
screen "4. VFD 10 - 13" 1280x800, template "Main_Template"
   on GenerateScreen: SetTag("animation_page", 4)
   Bar "Bar_1" at 206,213 size 88x440; MinimumValue 0; MaximumValue 50
      ProcessValue <- "speedActual_address_10"
   Button "Button_7" at 35,514 size 150x62; TextOff '+'
      on Press: function_b14e0dd5("increaseSpeed_address_10", 0)
      Appearance <- "statusIncrease_address_10"
   Button "Button_8" at 35,591 size 150x62; TextOff '-'
      on Press: function_b14e0dd5("decreaseSpeed_address_10", 0)
      Appearance <- "statusDecrease_address_10"
   TextField "Text field_20" at 35,428 size 150x62; Text 'Hz'
   IOField "I/O field_1" at 37,430 size 98x57; FormatPattern 99.99
      ProcessValue <- "speedActual_address_10"
   TextField "Text field_14" at 28,133 size 207x62; Text 'Gauge Roll 3rd Set'
   TextField "Text field_26" at 35,228 size 150x62; Text 'Hz'
   TextField "Text field_32" at 35,328 size 150x62; Text 'Hz'
   IOField "I/O field_2" at 39,231 size 98x57; FormatPattern 99.99
      ProcessValue <- "speedReff_singleSync_address_10"
   TextField "Text field_1" at 35,400 size 115x27; Text 'Actual Speed'
   TextField "Text field_2" at 35,302 size 144x27; Text 'Reff Speed Sync'
   TextField "Text field_3" at 35,200 size 155x27; Text 'Reff Speed Single'
   TextField "Text field_4" at 36,661 size 149x45; Text 'VFD 10'
      Appearance <- "Running_Motor Addres_10"
   Bar "Bar_2" at 518,213 size 88x440; MinimumValue 0; MaximumValue 50
      ProcessValue <- "speedActual_address_11"
   Button "Button_2" at 347,514 size 150x62; TextOff '+'
      on Press: function_b14e0dd5("increaseSpeed_address_11", 0)
      Appearance <- "statusIncrease_address_11"
   Button "Button_3" at 347,591 size 150x62; TextOff '-'
      on Press: function_b14e0dd5("decreaseSpeed_address_11", 0)
      Appearance <- "statusDecrease_address_11"
   TextField "Text field_5" at 347,428 size 150x62; Text 'Hz'
   IOField "I/O field_3" at 349,430 size 98x57; FormatPattern 99.99
      ProcessValue <- "speedActual_address_11"
   TextField "Text field_6" at 340,133 size 207x62; Text 'Conveyor of Gauge Roll 3rd Set'
   TextField "Text field_7" at 347,228 size 150x62; Text 'Hz'
   TextField "Text field_8" at 347,328 size 150x62; Text 'Hz'
   IOField "I/O field_4" at 351,231 size 98x57; FormatPattern 99.99
      ProcessValue <- "speedReff_singleSync_address_11"
   TextField "Text field_9" at 347,400 size 115x27; Text 'Actual Speed'
   TextField "Text field_10" at 347,302 size 144x27; Text 'Reff Speed Sync'
   TextField "Text field_11" at 347,200 size 155x27; Text 'Reff Speed Single'
   TextField "Text field_12" at 348,661 size 149x45; Text 'VFD 11'
      Appearance <- "Running_Motor Addres_11"
   Bar "Bar_3" at 830,213 size 88x440; MinimumValue 0; MaximumValue 50
      ProcessValue <- "speedActual_address_12"
   Button "Button_4" at 659,514 size 150x62; TextOff '+'
      on Press: function_b14e0dd5("increaseSpeed_address_12", 0)
      Appearance <- "statusIncrease_address_12"
   Button "Button_5" at 659,591 size 150x62; TextOff '-'
      on Press: function_b14e0dd5("decreaseSpeed_address_12", 0)
      Appearance <- "statusDecrease_address_12"
   TextField "Text field_13" at 659,428 size 150x62; Text 'Hz'
   IOField "I/O field_5" at 661,430 size 98x57; FormatPattern 99.99
      ProcessValue <- "speedActual_address_12"
   TextField "Text field_15" at 652,133 size 207x62; Text 'Passing Conveyor of Rotary Mould'
   TextField "Text field_16" at 659,228 size 150x62; Text 'Hz'
   TextField "Text field_17" at 659,328 size 150x62; Text 'Hz'
   IOField "I/O field_6" at 663,231 size 98x57; FormatPattern 99.99
      ProcessValue <- "speedReff_singleSync_address_12"
   TextField "Text field_18" at 659,400 size 115x27; Text 'Actual Speed'
   TextField "Text field_19" at 659,302 size 144x27; Text 'Reff Speed Sync'
   TextField "Text field_21" at 659,200 size 155x27; Text 'Reff Speed Single'
   TextField "Text field_22" at 660,661 size 149x45; Text 'VFD 12'
      Appearance <- "Running_Motor Addres_12"
   Bar "Bar_4" at 1142,213 size 88x440; MinimumValue 0; MaximumValue 50
      ProcessValue <- "speedActual_address_13"
   Button "Button_6" at 971,514 size 150x62; TextOff '+'
      on Press: function_b14e0dd5("increaseSpeed_address_13", 0)
      Appearance <- "statusIncrease_address_13"
   Button "Button_9" at 971,591 size 150x62; TextOff '-'
      on Press: function_b14e0dd5("decreaseSpeed_address_13", 0)
      Appearance <- "statusDecrease_address_13"
   TextField "Text field_23" at 971,428 size 150x62; Text 'Hz'
   IOField "I/O field_7" at 973,430 size 98x57; FormatPattern 99.99
      ProcessValue <- "speedActual_address_13"
   TextField "Text field_24" at 964,133 size 207x62; Text 'Conveyor of Rotary Moulder'
   TextField "Text field_25" at 971,228 size 150x62; Text 'Hz'
   TextField "Text field_27" at 971,328 size 150x62; Text 'Hz'
   IOField "I/O field_8" at 975,231 size 98x57; FormatPattern 99.99
      ProcessValue <- "speedReff_singleSync_address_13"
   TextField "Text field_28" at 971,400 size 115x27; Text 'Actual Speed'
   TextField "Text field_29" at 971,302 size 144x27; Text 'Reff Speed Sync'
   TextField "Text field_30" at 971,200 size 155x27; Text 'Reff Speed Single'
   TextField "Text field_31" at 972,661 size 149x45; Text 'VFD 13'
      Appearance <- "Running_Motor Addres_13"
   IOField "I/O field_14" at 349,330 size 98x57; FormatPattern 99.99
      ProcessValue <- "speedReff_NOT_singleSync_address_11"
   IOField "I/O field_9" at 661,330 size 98x57; FormatPattern 99.99
      ProcessValue <- "speedReff_NOT_singleSync_address_12"
   IOField "I/O field_10" at 973,330 size 98x57; FormatPattern 99.99
      ProcessValue <- "speedReff_NOT_singleSync_address_13"
   SymbolicIOField "Symbolic I/O field_2" at 550,133 size 77x62; TextOn '1'; TextOff '0'; TextList "Mode_Syncron"
      Appearance <- "Syncron_2"
      ProcessValue <- "Syncron_2"
   SymbolicIOField "Symbolic I/O field_3" at 862,133 size 77x62; TextOn '1'; TextOff '0'; TextList "Mode_Syncron"
      Appearance <- "Syncron_2"
      ProcessValue <- "Syncron_2"
   SymbolicIOField "Symbolic I/O field_4" at 1174,133 size 77x62; TextOn '1'; TextOff '0'; TextList "Mode_Syncron"
      Appearance <- "Syncron_1"
      ProcessValue <- "Syncron_1"
   IOField "I/O field_11" at 37,330 size 98x57; FormatPattern 99.99
      ProcessValue <- "speedReff_NOT_singleSync_address_10"
   SymbolicIOField "Symbolic I/O field_1" at 238,133 size 77x62; TextOn '1'; TextOff '0'; TextList "Mode_Syncron"
      Appearance <- "Syncron_2"
      ProcessValue <- "Syncron_2"
   Button "Button_1" at 0,721 size 160x79; TextOff 'MAIN'
      on Click: ActivateScreen("1. MAIN", 0)
      Appearance <- "animation_page"
   Button "Button_10" at 160,721 size 160x79; TextOff 'VFD 2 - 5'
      on Click: ActivateScreen("2. VFD 2 - 5", 0)
      Appearance <- "animation_page"
   Button "Button_11" at 320,721 size 160x79; TextOff 'VFD 6 - 9'
      on Click: ActivateScreen("3. VFD 6 - 9", 0)
      Appearance <- "animation_page"
   Button "Button_12" at 480,721 size 160x79; TextOff 'VFD 10 - 13'
      on Click: ActivateScreen("4. VFD 10 - 13", 0)
      Appearance <- "animation_page"
   Button "Button_13" at 640,721 size 160x79; TextOff 'VFD 14 - 17'
      on Click: ActivateScreen("5. VFD 14 - 17", 0)
      Appearance <- "animation_page"
   Button "Button_14" at 800,721 size 160x79; TextOff 'VFD 18 - 21'
      on Click: ActivateScreen("6. VFD 18 - 21", 0)
      Appearance <- "animation_page"
   Button "Button_15" at 960,721 size 160x79; TextOff 'VFD 22 - 23'
      on Click: ActivateScreen("7. VFD 22 - 23", 0)
      Appearance <- "animation_page"
   Button "Button_16" at 1120,721 size 160x79; TextOff 'Alarm'
      on Click: ActivateScreen("8. ALARM", 0)
      Appearance <- "animation_page"
   TextField "Text field_34" at 0,64 size 331x50; Text 'MOTOR CONTROL SPEED'
   Softkey "Softkey_F1" at 0,0 size 0x0
      on KeyDown: ActivateScreen("1. MAIN", 0)
   Softkey "Softkey_F2" at 0,0 size 0x0
      on KeyDown: ActivateScreen("2. VFD 2 - 5", 0)
   Softkey "Softkey_F3" at 0,0 size 0x0
      on KeyDown: ActivateScreen("3. VFD 6 - 9", 0)
   Softkey "Softkey_F4" at 0,0 size 0x0
      on KeyDown: ActivateScreen("4. VFD 10 - 13", 0)
   Softkey "Softkey_F5" at 0,0 size 0x0
      on KeyDown: ActivateScreen("5. VFD 14 - 17", 0)
   Softkey "Softkey_F6" at 0,0 size 0x0
      on KeyDown: ActivateScreen("6. VFD 18 - 21", 0)
   Softkey "Softkey_F7" at 0,0 size 0x0
      on KeyDown: ActivateScreen("7. VFD 22 - 23", 0)
   Softkey "Softkey_F8" at 0,0 size 0x0
      on KeyDown: ActivateScreen("8. ALARM", 0)
   Softkey "Softkey_F9" at 0,0 size 0x0
      on KeyDown: ActivateScreen("9. VFD PROFIBUS", 0)
   Softkey "Softkey_F10" at 0,0 size 0x0
      on KeyDown: ActivateScreen("10. SETTINGS", 0)

screen "5. VFD 14 - 17" 1280x800, template "Main_Template"
   on GenerateScreen: SetTag("animation_page", 5)
   Bar "Bar_1" at 206,213 size 88x440; MinimumValue 0; MaximumValue 50
      ProcessValue <- "speedActual_address_14"
   Button "Button_7" at 35,514 size 150x62; TextOff '+'
      on Press: function_b14e0dd5("increaseSpeed_address_14", 0)
      Appearance <- "statusIncrease_address_14"
   Button "Button_8" at 35,591 size 150x62; TextOff '-'
      on Press: function_b14e0dd5("decreaseSpeed_address_14", 0)
      Appearance <- "statusDecrease_address_14"
   TextField "Text field_20" at 35,428 size 150x62; Text 'Hz'
   IOField "I/O field_1" at 37,430 size 98x57; FormatPattern 99.99
      ProcessValue <- "speedActual_address_14"
   TextField "Text field_14" at 28,133 size 207x62; Text 'Drive of Mould'
   TextField "Text field_26" at 35,228 size 150x62; Text 'Hz'
   TextField "Text field_32" at 35,328 size 150x62; Text 'Hz'
   IOField "I/O field_2" at 39,231 size 98x57; FormatPattern 99.99
      ProcessValue <- "speedReff_singleSync_address_14"
   TextField "Text field_1" at 35,400 size 115x27; Text 'Actual Speed'
   TextField "Text field_2" at 35,302 size 144x27; Text 'Reff Speed Sync'
   TextField "Text field_3" at 35,200 size 155x27; Text 'Reff Speed Single'
   TextField "Text field_4" at 36,661 size 149x45; Text 'VFD 14'
      Appearance <- "Running_Motor Addres_14"
   Bar "Bar_2" at 518,213 size 88x440; MinimumValue 0; MaximumValue 50
      ProcessValue <- "speedActual_address_15"
   Button "Button_2" at 347,514 size 150x62; TextOff '+'
      on Press: function_b14e0dd5("increaseSpeed_address_15", 0)
      Appearance <- "statusIncrease_address_15"
   Button "Button_3" at 347,591 size 150x62; TextOff '-'
      on Press: function_b14e0dd5("decreaseSpeed_address_15", 0)
      Appearance <- "statusDecrease_address_15"
   TextField "Text field_5" at 347,428 size 150x62; Text 'Hz'
   IOField "I/O field_3" at 349,430 size 98x57; FormatPattern 99.99
      ProcessValue <- "speedActual_address_15"
   TextField "Text field_6" at 340,133 size 207x62; Text 'Forcing Roll'
   TextField "Text field_7" at 347,228 size 150x62; Text 'Hz'
   TextField "Text field_8" at 347,328 size 150x62; Text 'Hz'
   IOField "I/O field_4" at 351,231 size 98x57; FormatPattern 99.99
      ProcessValue <- "speedReff_singleSync_address_15"
   TextField "Text field_9" at 347,400 size 115x27; Text 'Actual Speed'
   TextField "Text field_10" at 347,302 size 144x27; Text 'Reff Speed Sync'
   TextField "Text field_11" at 347,200 size 155x27; Text 'Reff Speed Single'
   TextField "Text field_12" at 348,661 size 149x45; Text 'VFD 15'
      Appearance <- "Running_Motor Addres_15"
   Bar "Bar_3" at 830,213 size 88x440; MinimumValue 0; MaximumValue 50
      ProcessValue <- "speedActual_address_16"
   Button "Button_4" at 659,514 size 150x62; TextOff '+'
      on Press: function_b14e0dd5("increaseSpeed_address_16", 0)
      Appearance <- "statusIncrease_address_16"
   Button "Button_5" at 659,591 size 150x62; TextOff '-'
      on Press: function_b14e0dd5("decreaseSpeed_address_16", 0)
      Appearance <- "statusDecrease_address_16"
   TextField "Text field_13" at 659,428 size 150x62; Text 'Hz'
   IOField "I/O field_5" at 661,430 size 98x57; FormatPattern 99.99
      ProcessValue <- "speedActual_address_16"
   TextField "Text field_15" at 652,133 size 207x62; Text 'Mould of Rotary Cutter'
   TextField "Text field_16" at 659,228 size 150x62; Text 'Hz'
   TextField "Text field_17" at 659,328 size 150x62; Text 'Hz'
   IOField "I/O field_6" at 663,231 size 98x57; FormatPattern 99.99
      ProcessValue <- "speedReff_singleSync_address_16"
   TextField "Text field_18" at 659,400 size 115x27; Text 'Actual Speed'
   TextField "Text field_19" at 659,302 size 144x27; Text 'Reff Speed Sync'
   TextField "Text field_21" at 659,200 size 155x27; Text 'Reff Speed Single'
   TextField "Text field_22" at 660,661 size 149x45; Text 'VFD 16'
      Appearance <- "Running_Motor Addres_16"
   Bar "Bar_4" at 1142,213 size 88x440; MinimumValue 0; MaximumValue 50
      ProcessValue <- "speedActual_address_17"
   Button "Button_6" at 971,514 size 150x62; TextOff '+'
      on Press: function_b14e0dd5("increaseSpeed_address_17", 0)
      Appearance <- "statusIncrease_address_17"
   Button "Button_9" at 971,591 size 150x62; TextOff '-'
      on Press: function_b14e0dd5("decreaseSpeed_address_17", 0)
      Appearance <- "statusDecrease_address_17"
   TextField "Text field_23" at 971,428 size 150x62; Text 'Hz'
   IOField "I/O field_7" at 973,430 size 98x57; FormatPattern 99.99
      ProcessValue <- "speedActual_address_17"
   TextField "Text field_24" at 964,133 size 207x62; Text 'Conveyor for Rotary Cutter'
   TextField "Text field_25" at 971,228 size 150x62; Text 'Hz'
   TextField "Text field_27" at 971,328 size 150x62; Text 'Hz'
   IOField "I/O field_8" at 975,231 size 98x57; FormatPattern 99.99
      ProcessValue <- "speedReff_singleSync_address_17"
   TextField "Text field_28" at 971,400 size 115x27; Text 'Actual Speed'
   TextField "Text field_29" at 971,302 size 144x27; Text 'Reff Speed Sync'
   TextField "Text field_30" at 971,200 size 155x27; Text 'Reff Speed Single'
   TextField "Text field_31" at 972,661 size 149x45; Text 'VFD 17'
      Appearance <- "Running_Motor Addres_17"
   IOField "I/O field_14" at 349,330 size 98x57; FormatPattern 99.99
      ProcessValue <- "speedReff_NOT_singleSync_address_15"
   IOField "I/O field_9" at 661,330 size 98x57; FormatPattern 99.99
      ProcessValue <- "speedReff_NOT_singleSync_address_16"
   IOField "I/O field_10" at 973,330 size 98x57; FormatPattern 99.99
      ProcessValue <- "speedReff_NOT_singleSync_address_17"
   SymbolicIOField "Symbolic I/O field_2" at 550,133 size 77x62; TextOn '1'; TextOff '0'; TextList "Mode_Syncron"
      Appearance <- "Syncron_1"
      ProcessValue <- "Syncron_1"
   SymbolicIOField "Symbolic I/O field_3" at 862,133 size 77x62; TextOn '1'; TextOff '0'; TextList "Mode_Syncron"
      Appearance <- "Syncron_2"
      ProcessValue <- "Syncron_2"
   SymbolicIOField "Symbolic I/O field_4" at 1174,133 size 77x62; TextOn '1'; TextOff '0'; TextList "Mode_Syncron"
      Appearance <- "Syncron_3"
      ProcessValue <- "Syncron_3"
   IOField "I/O field_11" at 37,330 size 98x57; FormatPattern 99.99
      ProcessValue <- "speedReff_NOT_singleSync_address_14"
   SymbolicIOField "Symbolic I/O field_1" at 238,133 size 77x62; TextOn '1'; TextOff '0'; TextList "Mode_Syncron"
      Appearance <- "Syncron_1"
      ProcessValue <- "Syncron_1"
   Button "Button_1" at 0,721 size 160x79; TextOff 'MAIN'
      on Click: ActivateScreen("1. MAIN", 0)
      Appearance <- "animation_page"
   Button "Button_10" at 160,721 size 160x79; TextOff 'VFD 2 - 5'
      on Click: ActivateScreen("2. VFD 2 - 5", 0)
      Appearance <- "animation_page"
   Button "Button_11" at 320,721 size 160x79; TextOff 'VFD 6 - 9'
      on Click: ActivateScreen("3. VFD 6 - 9", 0)
      Appearance <- "animation_page"
   Button "Button_12" at 480,721 size 160x79; TextOff 'VFD 10 - 13'
      on Click: ActivateScreen("4. VFD 10 - 13", 0)
      Appearance <- "animation_page"
   Button "Button_13" at 640,721 size 160x79; TextOff 'VFD 14 - 17'
      on Click: ActivateScreen("5. VFD 14 - 17", 0)
      Appearance <- "animation_page"
   Button "Button_14" at 800,721 size 160x79; TextOff 'VFD 18 - 21'
      on Click: ActivateScreen("6. VFD 18 - 21", 0)
      Appearance <- "animation_page"
   Button "Button_15" at 960,721 size 160x79; TextOff 'VFD 22 - 23'
      on Click: ActivateScreen("7. VFD 22 - 23", 0)
      Appearance <- "animation_page"
   Button "Button_16" at 1120,721 size 160x79; TextOff 'Alarm'
      on Click: ActivateScreen("8. ALARM", 0)
      Appearance <- "animation_page"
   TextField "Text field_34" at 0,64 size 331x50; Text 'MOTOR CONTROL SPEED'
   Softkey "Softkey_F5" at 0,0 size 0x0
      on KeyDown: ActivateScreen("5. VFD 14 - 17", 0)
   Softkey "Softkey_F1" at 0,0 size 0x0
      on KeyDown: ActivateScreen("1. MAIN", 0)
   Softkey "Softkey_F2" at 0,0 size 0x0
      on KeyDown: ActivateScreen("2. VFD 2 - 5", 0)
   Softkey "Softkey_F3" at 0,0 size 0x0
      on KeyDown: ActivateScreen("3. VFD 6 - 9", 0)
   Softkey "Softkey_F4" at 0,0 size 0x0
      on KeyDown: ActivateScreen("4. VFD 10 - 13", 0)
   Softkey "Softkey_F6" at 0,0 size 0x0
      on KeyDown: ActivateScreen("6. VFD 18 - 21", 0)
   Softkey "Softkey_F7" at 0,0 size 0x0
      on KeyDown: ActivateScreen("7. VFD 22 - 23", 0)
   Softkey "Softkey_F8" at 0,0 size 0x0
      on KeyDown: ActivateScreen("8. ALARM", 0)
   Softkey "Softkey_F9" at 0,0 size 0x0
      on KeyDown: ActivateScreen("9. VFD PROFIBUS", 0)
   Softkey "Softkey_F10" at 0,0 size 0x0
      on KeyDown: ActivateScreen("10. SETTINGS", 0)

screen "6. VFD 18 - 21" 1280x800, template "Main_Template"
   on GenerateScreen: SetTag("animation_page", 6)
   Bar "Bar_1" at 206,213 size 88x440; MinimumValue 0; MaximumValue 50
      ProcessValue <- "speedActual_address_18"
   Button "Button_7" at 35,514 size 150x62; TextOff '+'
      on Press: function_b14e0dd5("increaseSpeed_address_18", 0)
      Appearance <- "statusIncrease_address_18"
   Button "Button_8" at 35,591 size 150x62; TextOff '-'
      on Press: function_b14e0dd5("decreaseSpeed_address_18", 0)
      Appearance <- "statusDecrease_address_18"
   TextField "Text field_20" at 35,428 size 150x62; Text 'Hz'
   IOField "I/O field_1" at 37,430 size 98x57; FormatPattern 99.99
      ProcessValue <- "speedActual_address_18"
   TextField "Text field_14" at 28,133 size 207x62; Text 'Dough Feed for Rotary Moulder'
   TextField "Text field_26" at 35,228 size 150x62; Text 'Hz'
   TextField "Text field_32" at 35,328 size 150x62; Text 'Hz'
   IOField "I/O field_2" at 39,231 size 98x57; FormatPattern 99.99
      ProcessValue <- "speedReff_singleSync_address_18"
   TextField "Text field_1" at 35,400 size 115x27; Text 'Actual Speed'
   TextField "Text field_2" at 35,302 size 144x27; Text 'Reff Speed Sync'
   TextField "Text field_3" at 35,200 size 155x27; Text 'Reff Speed Single'
   TextField "Text field_4" at 36,661 size 149x45; Text 'VFD 18'
      Appearance <- "Running_Motor Addres_18"
   Bar "Bar_2" at 518,213 size 88x440; MinimumValue 0; MaximumValue 50
      ProcessValue <- "speedActual_address_19"
   Button "Button_2" at 347,514 size 150x62; TextOff '+'
      on Press: function_b14e0dd5("increaseSpeed_address_19", 0)
      Appearance <- "statusIncrease_address_19"
   Button "Button_3" at 347,591 size 150x62; TextOff '-'
      on Press: function_b14e0dd5("decreaseSpeed_address_19", 0)
      Appearance <- "statusDecrease_address_19"
   TextField "Text field_5" at 347,428 size 150x62; Text 'Hz'
   IOField "I/O field_3" at 349,430 size 98x57; FormatPattern 99.99
      ProcessValue <- "speedActual_address_19"
   TextField "Text field_6" at 340,133 size 207x62; Text 'Conveyor of Scrapt Lift Passing'
   TextField "Text field_7" at 347,228 size 150x62; Text 'Hz'
   TextField "Text field_8" at 347,328 size 150x62; Text 'Hz'
   IOField "I/O field_4" at 351,231 size 98x57; FormatPattern 99.99
      ProcessValue <- "speedReff_singleSync_address_19"
   TextField "Text field_9" at 347,400 size 115x27; Text 'Actual Speed'
   TextField "Text field_10" at 347,302 size 144x27; Text 'Reff Speed Sync'
   TextField "Text field_11" at 347,200 size 155x27; Text 'Reff Speed Single'
   TextField "Text field_12" at 348,661 size 149x45; Text 'VFD 19'
      Appearance <- "Running_Motor Addres_19"
   Bar "Bar_3" at 830,213 size 88x440; MinimumValue 0; MaximumValue 50
      ProcessValue <- "speedActual_address_20"
   Button "Button_4" at 659,514 size 150x62; TextOff '+'
      on Press: function_b14e0dd5("increaseSpeed_address_20", 0)
      Appearance <- "statusIncrease_address_20"
   Button "Button_5" at 659,591 size 150x62; TextOff '-'
      on Press: function_b14e0dd5("decreaseSpeed_address_20", 0)
      Appearance <- "statusDecrease_address_20"
   TextField "Text field_13" at 659,428 size 150x62; Text 'Hz'
   IOField "I/O field_5" at 661,430 size 98x57; FormatPattern 99.99
      ProcessValue <- "speedActual_address_20"
   TextField "Text field_15" at 652,133 size 207x62; Text 'Conveyor of Salt Sprinkler'
   TextField "Text field_16" at 659,228 size 150x62; Text 'Hz'
   TextField "Text field_17" at 659,328 size 150x62; Text 'Hz'
   IOField "I/O field_6" at 663,231 size 98x57; FormatPattern 99.99
      ProcessValue <- "speedReff_singleSync_address_20"
   TextField "Text field_18" at 659,400 size 115x27; Text 'Actual Speed'
   TextField "Text field_19" at 659,302 size 144x27; Text 'Reff Speed Sync'
   TextField "Text field_21" at 659,200 size 155x27; Text 'Reff Speed Single'
   TextField "Text field_22" at 660,661 size 149x45; Text 'VFD 20'
      Appearance <- "Running_Motor Addres_20"
   Bar "Bar_4" at 1142,213 size 88x440; MinimumValue 0; MaximumValue 50
      ProcessValue <- "speedActual_address_21"
   Button "Button_6" at 971,514 size 150x62; TextOff '+'
      on Press: function_b14e0dd5("increaseSpeed_address_21", 0)
      Appearance <- "statusIncrease_address_21"
   Button "Button_9" at 971,591 size 150x62; TextOff '-'
      on Press: function_b14e0dd5("decreaseSpeed_address_21", 0)
      Appearance <- "statusDecrease_address_21"
   TextField "Text field_23" at 971,428 size 150x62; Text 'Hz'
   IOField "I/O field_7" at 973,430 size 98x57; FormatPattern 99.99
      ProcessValue <- "speedActual_address_21"
   TextField "Text field_24" at 964,133 size 207x62; Text 'Recovery Conveyor of Salt Sprinkler'
   TextField "Text field_25" at 971,228 size 150x62; Text 'Hz'
   TextField "Text field_27" at 971,328 size 150x62; Text 'Hz'
   IOField "I/O field_8" at 975,231 size 98x57; FormatPattern 99.99
      ProcessValue <- "speedReff_singleSync_address_21"
   TextField "Text field_28" at 971,400 size 115x27; Text 'Actual Speed'
   TextField "Text field_29" at 971,302 size 144x27; Text 'Reff Speed Sync'
   TextField "Text field_30" at 971,200 size 155x27; Text 'Reff Speed Single'
   TextField "Text field_31" at 972,661 size 149x45; Text 'VFD 21'
      Appearance <- "Running_Motor Addres_21"
   IOField "I/O field_14" at 349,330 size 98x57; FormatPattern 99.99
      ProcessValue <- "speedReff_NOT_singleSync_address_19"
   IOField "I/O field_9" at 661,330 size 98x57; FormatPattern 99.99
      ProcessValue <- "speedReff_NOT_singleSync_address_20"
   IOField "I/O field_10" at 973,330 size 98x57; FormatPattern 99.99
      ProcessValue <- "speedReff_NOT_singleSync_address_21"
   SymbolicIOField "Symbolic I/O field_2" at 550,133 size 77x62; TextOn '1'; TextOff '0'; TextList "Mode_Syncron"
      Appearance <- "Syncron_3"
      ProcessValue <- "Syncron_3"
   SymbolicIOField "Symbolic I/O field_4" at 1174,133 size 77x62; TextOn '1'; TextOff '0'; TextList "Mode_Syncron"
      Appearance <- "Syncron_3"
      ProcessValue <- "Syncron_3"
   IOField "I/O field_11" at 37,330 size 98x57; FormatPattern 99.99
      ProcessValue <- "speedReff_NOT_singleSync_address_18"
   TextField "Text field_33" at 238,133 size 76x62; Text 'Single'
   TextField "Text field_35" at 863,133 size 76x62; Text 'Single'
   Button "Button_1" at 0,721 size 160x79; TextOff 'MAIN'
      on Click: ActivateScreen("1. MAIN", 0)
      Appearance <- "animation_page"
   Button "Button_10" at 160,721 size 160x79; TextOff 'VFD 2 - 5'
      on Click: ActivateScreen("2. VFD 2 - 5", 0)
      Appearance <- "animation_page"
   Button "Button_11" at 320,721 size 160x79; TextOff 'VFD 6 - 9'
      on Click: ActivateScreen("3. VFD 6 - 9", 0)
      Appearance <- "animation_page"
   Button "Button_12" at 480,721 size 160x79; TextOff 'VFD 10 - 13'
      on Click: ActivateScreen("4. VFD 10 - 13", 0)
      Appearance <- "animation_page"
   Button "Button_13" at 640,721 size 160x79; TextOff 'VFD 14 - 17'
      on Click: ActivateScreen("5. VFD 14 - 17", 0)
      Appearance <- "animation_page"
   Button "Button_14" at 800,721 size 160x79; TextOff 'VFD 18 - 21'
      on Click: ActivateScreen("6. VFD 18 - 21", 0)
      Appearance <- "animation_page"
   Button "Button_15" at 960,721 size 160x79; TextOff 'VFD 22 - 23'
      on Click: ActivateScreen("7. VFD 22 - 23", 0)
      Appearance <- "animation_page"
   Button "Button_16" at 1120,721 size 160x79; TextOff 'Alarm'
      on Click: ActivateScreen("8. ALARM", 0)
      Appearance <- "animation_page"
   TextField "Text field_34" at 0,64 size 331x50; Text 'MOTOR CONTROL SPEED'
   Softkey "Softkey_F5" at 0,0 size 0x0
      on KeyDown: ActivateScreen("5. VFD 14 - 17", 0)
   Softkey "Softkey_F1" at 0,0 size 0x0
      on KeyDown: ActivateScreen("1. MAIN", 0)
   Softkey "Softkey_F2" at 0,0 size 0x0
      on KeyDown: ActivateScreen("2. VFD 2 - 5", 0)
   Softkey "Softkey_F3" at 0,0 size 0x0
      on KeyDown: ActivateScreen("3. VFD 6 - 9", 0)
   Softkey "Softkey_F4" at 0,0 size 0x0
      on KeyDown: ActivateScreen("4. VFD 10 - 13", 0)
   Softkey "Softkey_F6" at 0,0 size 0x0
      on KeyDown: ActivateScreen("6. VFD 18 - 21", 0)
   Softkey "Softkey_F7" at 0,0 size 0x0
      on KeyDown: ActivateScreen("7. VFD 22 - 23", 0)
   Softkey "Softkey_F8" at 0,0 size 0x0
      on KeyDown: ActivateScreen("8. ALARM", 0)
   Softkey "Softkey_F9" at 0,0 size 0x0
      on KeyDown: ActivateScreen("9. VFD PROFIBUS", 0)
   Softkey "Softkey_F10" at 0,0 size 0x0
      on KeyDown: ActivateScreen("10. SETTINGS", 0)

screen "7. VFD 22 - 23" 1280x800, template "Main_Template"
   on GenerateScreen: SetTag("animation_page", 7)
   Bar "Bar_1" at 206,213 size 88x440; MinimumValue 0; MaximumValue 50
      ProcessValue <- "speedActual_address_22"
   Button "Button_7" at 35,514 size 150x62; TextOff '+'
      on Press: function_b14e0dd5("increaseSpeed_address_22", 0)
      Appearance <- "statusIncrease_address_22"
   Button "Button_8" at 35,591 size 150x62; TextOff '-'
      on Press: function_b14e0dd5("decreaseSpeed_address_22", 0)
      Appearance <- "statusDecrease_address_22"
   TextField "Text field_20" at 35,428 size 150x62; Text 'Hz'
   IOField "I/O field_1" at 37,430 size 98x57; FormatPattern 99.99
      ProcessValue <- "speedActual_address_22"
   TextField "Text field_14" at 28,133 size 207x62; Text 'Conveyor Swivel Panner'
   TextField "Text field_26" at 35,228 size 150x62; Text 'Hz'
   TextField "Text field_32" at 35,328 size 150x62; Text 'Hz'
   IOField "I/O field_2" at 39,231 size 98x57; FormatPattern 99.99
      ProcessValue <- "speedReff_singleSync_address_22"
   TextField "Text field_1" at 35,400 size 115x27; Text 'Actual Speed'
   TextField "Text field_2" at 35,302 size 144x27; Text 'Reff Speed Sync'
   TextField "Text field_3" at 35,200 size 155x27; Text 'Reff Speed Single'
   TextField "Text field_4" at 36,661 size 149x45; Text 'VFD 22'
      Appearance <- "Running_Motor Addres_22"
   Bar "Bar_2" at 518,213 size 88x440; MinimumValue 0; MaximumValue 50
      ProcessValue <- "speedActual_address_23"
   Button "Button_2" at 347,514 size 150x62; TextOff '+'
      on Press: function_b14e0dd5("increaseSpeed_address_23", 0)
      Appearance <- "statusIncrease_address_23"
   Button "Button_3" at 347,591 size 150x62; TextOff '-'
      on Press: function_b14e0dd5("decreaseSpeed_address_23", 0)
      Appearance <- "statusDecrease_address_23"
   TextField "Text field_5" at 347,428 size 150x62; Text 'Hz'
   IOField "I/O field_3" at 349,430 size 98x57; FormatPattern 99.99
      ProcessValue <- "speedActual_address_23"
   TextField "Text field_6" at 340,133 size 207x62; Text 'Side Return VFD 23 for 4 Motor'
   TextField "Text field_7" at 347,228 size 150x62; Text 'Hz'
   TextField "Text field_8" at 347,328 size 150x62; Text 'Hz'
   IOField "I/O field_4" at 351,231 size 98x57; FormatPattern 99.99
      ProcessValue <- "speedReff_singleSync_address_23"
   TextField "Text field_9" at 347,400 size 115x27; Text 'Actual Speed'
   TextField "Text field_10" at 347,302 size 144x27; Text 'Reff Speed Sync'
   TextField "Text field_11" at 347,200 size 155x27; Text 'Reff Speed Single'
   TextField "Text field_12" at 348,661 size 149x45; Text 'VFD 23'
      Appearance <- "Running_Motor Addres_23"
   IOField "I/O field_14" at 349,330 size 98x57; FormatPattern 99.99
      ProcessValue <- "speedReff_NOT_singleSync_address_23"
   SymbolicIOField "Symbolic I/O field_2" at 550,133 size 77x62; TextOn '1'; TextOff '0'; TextList "Mode_Syncron"
      ProcessValue <- "Syncron_2"
      Appearance <- "Syncron_2"
   IOField "I/O field_11" at 37,330 size 98x57; FormatPattern 99.99
      ProcessValue <- "speedReff_NOT_singleSync_address_22"
   SymbolicIOField "Symbolic I/O field_1" at 238,133 size 77x62; TextOn '1'; TextOff '0'; TextList "Mode_Syncron"
      ProcessValue <- "Syncron_3"
      Appearance <- "Syncron_3"
   TextField "Text field_13" at 654,133 size 582x62; Text 'Menu'
   Button "Button_4" at 735,289 size 420x79; TextOff 'Communication Profibus'
      on Click: ActivateScreen("9. VFD PROFIBUS", 0)
   Button "Button_5" at 735,401 size 420x79; TextOff 'Diagnostic buffer view'
      on Click: ActivateScreen("11. DIAG", 0)
   Button "Button_6" at 735,513 size 420x79; TextOff 'Settings'
      on Click: ActivateScreen("10. SETTINGS", 0)
   TextField "Text field_34" at 0,64 size 331x50; Text 'MOTOR CONTROL SPEED'
   Button "Button_1" at 0,721 size 160x79; TextOff 'MAIN'
      on Click: ActivateScreen("1. MAIN", 0)
      Appearance <- "animation_page"
   Button "Button_10" at 160,721 size 160x79; TextOff 'VFD 2 - 5'
      on Click: ActivateScreen("2. VFD 2 - 5", 0)
      Appearance <- "animation_page"
   Button "Button_11" at 320,721 size 160x79; TextOff 'VFD 6 - 9'
      on Click: ActivateScreen("3. VFD 6 - 9", 0)
      Appearance <- "animation_page"
   Button "Button_12" at 480,721 size 160x79; TextOff 'VFD 10 - 13'
      on Click: ActivateScreen("4. VFD 10 - 13", 0)
      Appearance <- "animation_page"
   Button "Button_13" at 640,721 size 160x79; TextOff 'VFD 14 - 17'
      on Click: ActivateScreen("5. VFD 14 - 17", 0)
      Appearance <- "animation_page"
   Button "Button_14" at 800,721 size 160x79; TextOff 'VFD 18 - 21'
      on Click: ActivateScreen("6. VFD 18 - 21", 0)
      Appearance <- "animation_page"
   Button "Button_15" at 960,721 size 160x79; TextOff 'VFD 22 - 23'
      on Click: ActivateScreen("7. VFD 22 - 23", 0)
      Appearance <- "animation_page"
   Button "Button_16" at 1120,721 size 160x79; TextOff 'Alarm'
      on Click: ActivateScreen("8. ALARM", 0)
      Appearance <- "animation_page"
   Softkey "Softkey_F5" at 0,0 size 0x0
      on KeyDown: ActivateScreen("5. VFD 14 - 17", 0)
   Softkey "Softkey_F1" at 0,0 size 0x0
      on KeyDown: ActivateScreen("1. MAIN", 0)
   Softkey "Softkey_F2" at 0,0 size 0x0
      on KeyDown: ActivateScreen("2. VFD 2 - 5", 0)
   Softkey "Softkey_F3" at 0,0 size 0x0
      on KeyDown: ActivateScreen("3. VFD 6 - 9", 0)
   Softkey "Softkey_F4" at 0,0 size 0x0
      on KeyDown: ActivateScreen("4. VFD 10 - 13", 0)
   Softkey "Softkey_F6" at 0,0 size 0x0
      on KeyDown: ActivateScreen("6. VFD 18 - 21", 0)
   Softkey "Softkey_F7" at 0,0 size 0x0
      on KeyDown: ActivateScreen("7. VFD 22 - 23", 0)
   Softkey "Softkey_F8" at 0,0 size 0x0
      on KeyDown: ActivateScreen("8. ALARM", 0)
   Softkey "Softkey_F9" at 0,0 size 0x0
      on KeyDown: ActivateScreen("9. VFD PROFIBUS", 0)
   Softkey "Softkey_F10" at 0,0 size 0x0
      on KeyDown: ActivateScreen("10. SETTINGS", 0)

screen "12. DI/DO" 1280x800, template "Main_Template"
   Circle "Circle_1" at 551,250 size 23x23
      Appearance <- "In_124_0"
   Circle "Circle_2" at 551,274 size 23x23
      Appearance <- "In_124_1"
   Circle "Circle_3" at 551,298 size 23x23
      Appearance <- "In_124_2"
   Circle "Circle_4" at 551,322 size 23x23
      Appearance <- "In_124_3"
   Circle "Circle_5" at 551,346 size 23x23
      Appearance <- "In_124_4"
   Circle "Circle_6" at 551,370 size 23x23
      Appearance <- "In_124_5"
   Circle "Circle_7" at 551,394 size 23x23
      Appearance <- "In_124_6"
   Circle "Circle_8" at 551,418 size 23x23
      Appearance <- "In_124_7"
   Circle "Circle_9" at 551,467 size 23x23
      Appearance <- "In_125_0"
   Circle "Circle_10" at 551,491 size 23x23
      Appearance <- "In_125_1"
   Circle "Circle_11" at 551,515 size 23x23
      Appearance <- "In_125_2"
   Circle "Circle_12" at 551,539 size 23x23
      Appearance <- "In_125_3"
   Circle "Circle_13" at 551,563 size 23x23
      Appearance <- "In_125_4"
   Circle "Circle_14" at 551,587 size 23x23
      Appearance <- "In_125_5"
   Circle "Circle_15" at 551,611 size 23x23
      Appearance <- "In_125_6"
   Circle "Circle_16" at 551,635 size 23x23
      Appearance <- "In_125_7"
   Circle "Circle_17" at 623,250 size 23x23
      Appearance <- "In_126_0"
   Circle "Circle_18" at 623,274 size 23x23
      Appearance <- "In_126_1"
   Circle "Circle_19" at 623,298 size 23x23
      Appearance <- "In_126_2"
   Circle "Circle_20" at 623,322 size 23x23
      Appearance <- "In_126_3"
   Circle "Circle_21" at 623,346 size 23x23
      Appearance <- "In_126_4"
   Circle "Circle_22" at 623,370 size 23x23
      Appearance <- "In_126_5"
   Circle "Circle_23" at 623,394 size 23x23
      Appearance <- "In_126_6"
   Circle "Circle_24" at 623,418 size 23x23
      Appearance <- "In_126_7"
   Circle "Circle_25" at 623,467 size 23x23
      Appearance <- "In_127_0"
   Circle "Circle_26" at 623,491 size 23x23
      Appearance <- "In_127_1"
   Circle "Circle_27" at 623,515 size 23x23
      Appearance <- "In_127_2"
   Circle "Circle_28" at 623,539 size 23x23
      Appearance <- "In_127_3"
   Circle "Circle_29" at 623,563 size 23x23
      Appearance <- "In_127_4"
   Circle "Circle_30" at 623,587 size 23x23
      Appearance <- "In_127_5"
   Circle "Circle_31" at 623,611 size 23x23
      Appearance <- "In_127_6"
   Circle "Circle_32" at 623,635 size 23x23
      Appearance <- "In_127_7"
   Circle "Circle_33" at 697,250 size 23x23
      Appearance <- "Out_124_0"
   Circle "Circle_34" at 697,274 size 23x23
      Appearance <- "Out_124_1"
   Circle "Circle_35" at 697,298 size 23x23
      Appearance <- "Out_124_2"
   Circle "Circle_36" at 697,322 size 23x23
      Appearance <- "Out_124_3"
   Circle "Circle_37" at 697,346 size 23x23
      Appearance <- "Out_124_4"
   Circle "Circle_38" at 697,370 size 23x23
      Appearance <- "Out_124_5"
   Circle "Circle_39" at 697,394 size 23x23
      Appearance <- "Out_124_6"
   Circle "Circle_40" at 697,418 size 23x23
      Appearance <- "Out_124_7"
   Circle "Circle_41" at 697,467 size 23x23
      Appearance <- "Out_125_0"
   Circle "Circle_42" at 697,491 size 23x23
      Appearance <- "Out_125_1"
   Circle "Circle_43" at 697,515 size 23x23
      Appearance <- "Out_125_2"
   Circle "Circle_44" at 697,539 size 23x23
      Appearance <- "Out_125_3"
   Circle "Circle_45" at 697,563 size 23x23
      Appearance <- "Out_125_4"
   Circle "Circle_46" at 697,587 size 23x23
      Appearance <- "Out_125_5"
   Circle "Circle_47" at 697,611 size 23x23
      Appearance <- "Out_125_6"
   Circle "Circle_48" at 697,635 size 23x23
      Appearance <- "Out_125_7"
   Circle "Circle_49" at 807,250 size 23x23
      Appearance <- "In_0_0"
   Circle "Circle_50" at 807,274 size 23x23
      Appearance <- "In_0_1"
   Circle "Circle_51" at 807,298 size 23x23
      Appearance <- "In_0_2"
   Circle "Circle_52" at 807,322 size 23x23
      Appearance <- "In_0_3"
   Circle "Circle_53" at 807,346 size 23x23
      Appearance <- "In_0_4"
   Circle "Circle_54" at 807,370 size 23x23
      Appearance <- "In_0_5"
   Circle "Circle_55" at 807,394 size 23x23
      Appearance <- "In_0_6"
   Circle "Circle_56" at 807,418 size 23x23
      Appearance <- "In_0_7"
   Circle "Circle_57" at 807,467 size 23x23
      Appearance <- "In_1_0"
   Circle "Circle_58" at 807,491 size 23x23
      Appearance <- "In_1_1"
   Circle "Circle_59" at 807,515 size 23x23
      Appearance <- "In_1_2"
   Circle "Circle_60" at 807,539 size 23x23
      Appearance <- "In_1_3"
   Circle "Circle_61" at 807,563 size 23x23
      Appearance <- "In_1_4"
   Circle "Circle_62" at 807,587 size 23x23
      Appearance <- "In_1_5"
   Circle "Circle_63" at 807,611 size 23x23
      Appearance <- "In_1_6"
   Circle "Circle_64" at 807,635 size 23x23
      Appearance <- "In_1_7"
   Circle "Circle_65" at 879,250 size 23x23
      Appearance <- "In_2_0"
   Circle "Circle_66" at 879,274 size 23x23
      Appearance <- "In_2_1"
   Circle "Circle_67" at 879,298 size 23x23
      Appearance <- "In_2_2"
   Circle "Circle_68" at 879,322 size 23x23
      Appearance <- "In_2_3"
   Circle "Circle_69" at 879,346 size 23x23
      Appearance <- "In_2_4"
   Circle "Circle_70" at 879,370 size 23x23
      Appearance <- "In_2_5"
   Circle "Circle_71" at 879,394 size 23x23
      Appearance <- "In_2_6"
   Circle "Circle_72" at 879,418 size 23x23
      Appearance <- "In_2_7"
   Circle "Circle_73" at 879,467 size 23x23
      Appearance <- "In_3_0"
   Circle "Circle_74" at 879,491 size 23x23
      Appearance <- "In_3_1"
   Circle "Circle_75" at 879,515 size 23x23
      Appearance <- "In_3_2"
   Circle "Circle_76" at 879,539 size 23x23
      Appearance <- "In_3_3"
   Circle "Circle_77" at 879,563 size 23x23
      Appearance <- "In_3_4"
   Circle "Circle_78" at 879,587 size 23x23
      Appearance <- "In_3_5"
   Circle "Circle_79" at 879,611 size 23x23
      Appearance <- "In_3_6"
   Circle "Circle_80" at 879,635 size 23x23
      Appearance <- "In_3_7"
   Circle "Circle_81" at 935,250 size 23x23
      Appearance <- "In_4_0"
   Circle "Circle_82" at 935,274 size 23x23
      Appearance <- "In_4_1"
   Circle "Circle_83" at 935,298 size 23x23
      Appearance <- "In_4_2"
   Circle "Circle_84" at 935,322 size 23x23
      Appearance <- "In_4_3"
   Circle "Circle_85" at 935,346 size 23x23
      Appearance <- "In_4_4"
   Circle "Circle_86" at 935,370 size 23x23
      Appearance <- "In_4_5"
   Circle "Circle_87" at 935,394 size 23x23
      Appearance <- "In_4_6"
   Circle "Circle_88" at 935,418 size 23x23
      Appearance <- "In_4_7"
   Circle "Circle_89" at 935,467 size 23x23
      Appearance <- "In_5_0"
   Circle "Circle_90" at 935,491 size 23x23
      Appearance <- "In_5_1"
   Circle "Circle_91" at 935,515 size 23x23
      Appearance <- "In_5_2"
   Circle "Circle_92" at 935,539 size 23x23
      Appearance <- "In_5_3"
   Circle "Circle_93" at 935,563 size 23x23
      Appearance <- "In_5_4"
   Circle "Circle_94" at 935,587 size 23x23
      Appearance <- "In_5_5"
   Circle "Circle_95" at 935,611 size 23x23
      Appearance <- "In_5_6"
   Circle "Circle_96" at 935,635 size 23x23
      Appearance <- "In_5_7"
   Circle "Circle_97" at 1007,250 size 23x23
      Appearance <- "In_6_0"
   Circle "Circle_98" at 1007,274 size 23x23
      Appearance <- "In_6_1"
   Circle "Circle_99" at 1007,298 size 23x23
      Appearance <- "In_6_2"
   Circle "Circle_100" at 1007,322 size 23x23
      Appearance <- "In_6_3"
   Circle "Circle_101" at 1007,346 size 23x23
      Appearance <- "In_6_4"
   Circle "Circle_102" at 1007,370 size 23x23
      Appearance <- "In_6_5"
   Circle "Circle_103" at 1007,394 size 23x23
      Appearance <- "In_6_6"
   Circle "Circle_104" at 1007,418 size 23x23
      Appearance <- "In_6_7"
   Circle "Circle_105" at 1007,467 size 23x23
      Appearance <- "In_7_0"
   Circle "Circle_106" at 1007,491 size 23x23
      Appearance <- "In_7_1"
   Circle "Circle_107" at 1007,515 size 23x23
      Appearance <- "In_7_2"
   Circle "Circle_108" at 1007,539 size 23x23
      Appearance <- "In_7_3"
   Circle "Circle_109" at 1007,563 size 23x23
      Appearance <- "In_7_4"
   Circle "Circle_110" at 1007,587 size 23x23
      Appearance <- "In_7_5"
   Circle "Circle_111" at 1007,611 size 23x23
      Appearance <- "In_7_6"
   Circle "Circle_112" at 1007,635 size 23x23
      Appearance <- "In_7_7"
   TextField "Text field_38" at 0,64 size 331x50; Text 'SYSTEM DIAGNOSTIC / DI / DO'
   TextField "Text field_1" at 541,201 size 108x23; Text 'Digital Input'
   TextField "Text field_2" at 667,201 size 120x23; Text 'Digital Output'
   TextField "Text field_3" at 797,201 size 108x23; Text 'Digital Input'
   TextField "Text field_4" at 925,201 size 108x23; Text 'Digital Input'
   TextField "Text field_5" at 439,201 size 64x42; Text 'Comm Module'
   TextField "Text field_6" at 321,201 size 43x23; Text 'CPU'
   TextField "Text field_7" at 541,223 size 43x23; Text '124'
   TextField "Text field_8" at 541,447 size 43x23; Text '125'
   TextField "Text field_9" at 613,223 size 43x23; Text '126'
   TextField "Text field_10" at 687,223 size 43x23; Text '124'
   TextField "Text field_11" at 613,447 size 43x23; Text '127'
   TextField "Text field_12" at 575,248 size 33x20; Text '.0'
   TextField "Text field_13" at 575,272 size 33x20; Text '.1'
   TextField "Text field_14" at 575,296 size 33x20; Text '.2'
   TextField "Text field_15" at 575,320 size 33x20; Text '.3'
   TextField "Text field_16" at 575,344 size 33x20; Text '.4'
   TextField "Text field_17" at 575,368 size 33x20; Text '.5'
   TextField "Text field_18" at 575,392 size 33x20; Text '.6'
   TextField "Text field_19" at 575,416 size 33x20; Text '.7'
   TextField "Text field_20" at 602,248 size 33x20; Text '.0'
   TextField "Text field_21" at 602,272 size 33x20; Text '.1'
   TextField "Text field_22" at 602,296 size 33x20; Text '.2'
   TextField "Text field_23" at 602,320 size 33x20; Text '.3'
   TextField "Text field_24" at 602,344 size 33x20; Text '.4'
   TextField "Text field_25" at 602,368 size 33x20; Text '.5'
   TextField "Text field_26" at 602,392 size 33x20; Text '.6'
   TextField "Text field_27" at 602,416 size 33x20; Text '.7'
   TextField "Text field_28" at 723,248 size 33x20; Text '.0'
   TextField "Text field_29" at 723,272 size 33x20; Text '.1'
   TextField "Text field_30" at 723,296 size 33x20; Text '.2'
   TextField "Text field_31" at 723,320 size 33x20; Text '.3'
   TextField "Text field_32" at 723,344 size 33x20; Text '.4'
   TextField "Text field_33" at 723,368 size 33x20; Text '.5'
   TextField "Text field_34" at 723,392 size 33x20; Text '.6'
   TextField "Text field_35" at 723,416 size 33x20; Text '.7'
   TextField "Text field_36" at 831,248 size 33x20; Text '.0'
   TextField "Text field_37" at 831,272 size 33x20; Text '.1'
   TextField "Text field_39" at 831,296 size 33x20; Text '.2'
   TextField "Text field_40" at 831,320 size 33x20; Text '.3'
   TextField "Text field_41" at 831,344 size 33x20; Text '.4'
   TextField "Text field_42" at 831,368 size 33x20; Text '.5'
   TextField "Text field_43" at 831,392 size 33x20; Text '.6'
   TextField "Text field_44" at 831,416 size 33x20; Text '.7'
   TextField "Text field_45" at 959,248 size 33x20; Text '.0'
   TextField "Text field_46" at 959,272 size 33x20; Text '.1'
   TextField "Text field_47" at 959,296 size 33x20; Text '.2'
   TextField "Text field_48" at 959,320 size 33x20; Text '.3'
   TextField "Text field_49" at 959,344 size 33x20; Text '.4'
   TextField "Text field_50" at 959,368 size 33x20; Text '.5'
   TextField "Text field_51" at 959,392 size 33x20; Text '.6'
   TextField "Text field_52" at 959,416 size 33x20; Text '.7'
   TextField "Text field_53" at 986,248 size 33x20; Text '.0'
   TextField "Text field_54" at 986,272 size 33x20; Text '.1'
   TextField "Text field_55" at 986,296 size 33x20; Text '.2'
   TextField "Text field_56" at 986,320 size 33x20; Text '.3'
   TextField "Text field_57" at 986,344 size 33x20; Text '.4'
   TextField "Text field_58" at 986,368 size 33x20; Text '.5'
   TextField "Text field_59" at 986,392 size 33x20; Text '.6'
   TextField "Text field_60" at 986,416 size 33x20; Text '.7'
   TextField "Text field_61" at 858,248 size 33x20; Text '.0'
   TextField "Text field_62" at 858,272 size 33x20; Text '.1'
   TextField "Text field_63" at 858,296 size 33x20; Text '.2'
   TextField "Text field_64" at 858,320 size 33x20; Text '.3'
   TextField "Text field_65" at 858,344 size 33x20; Text '.4'
   TextField "Text field_66" at 858,368 size 33x20; Text '.5'
   TextField "Text field_67" at 858,392 size 33x20; Text '.6'
   TextField "Text field_68" at 858,416 size 33x20; Text '.7'
   TextField "Text field_69" at 575,467 size 33x20; Text '.0'
   TextField "Text field_70" at 575,491 size 33x20; Text '.1'
   TextField "Text field_71" at 575,515 size 33x20; Text '.2'
   TextField "Text field_72" at 575,539 size 33x20; Text '.3'
   TextField "Text field_73" at 575,563 size 33x20; Text '.4'
   TextField "Text field_74" at 575,587 size 33x20; Text '.5'
   TextField "Text field_75" at 575,611 size 33x20; Text '.6'
   TextField "Text field_76" at 575,635 size 33x20; Text '.7'
   TextField "Text field_77" at 602,467 size 33x20; Text '.0'
   TextField "Text field_78" at 602,491 size 33x20; Text '.1'
   TextField "Text field_79" at 602,515 size 33x20; Text '.2'
   TextField "Text field_80" at 602,539 size 33x20; Text '.3'
   TextField "Text field_81" at 602,563 size 33x20; Text '.4'
   TextField "Text field_82" at 602,587 size 33x20; Text '.5'
   TextField "Text field_83" at 602,611 size 33x20; Text '.6'
   TextField "Text field_84" at 602,635 size 33x20; Text '.7'
   TextField "Text field_85" at 723,467 size 33x20; Text '.0'
   TextField "Text field_86" at 723,491 size 33x20; Text '.1'
   TextField "Text field_87" at 723,515 size 33x20; Text '.2'
   TextField "Text field_88" at 723,539 size 33x20; Text '.3'
   TextField "Text field_89" at 723,563 size 33x20; Text '.4'
   TextField "Text field_90" at 723,587 size 33x20; Text '.5'
   TextField "Text field_91" at 723,611 size 33x20; Text '.6'
   TextField "Text field_92" at 723,635 size 33x20; Text '.7'
   TextField "Text field_93" at 831,467 size 33x20; Text '.0'
   TextField "Text field_94" at 831,491 size 33x20; Text '.1'
   TextField "Text field_95" at 831,515 size 33x20; Text '.2'
   TextField "Text field_96" at 831,539 size 33x20; Text '.3'
   TextField "Text field_97" at 831,563 size 33x20; Text '.4'
   TextField "Text field_98" at 831,587 size 33x20; Text '.5'
   TextField "Text field_99" at 831,611 size 33x20; Text '.6'
   TextField "Text field_100" at 831,635 size 33x20; Text '.7'
   TextField "Text field_101" at 959,467 size 33x20; Text '.0'
   TextField "Text field_102" at 959,491 size 33x20; Text '.1'
   TextField "Text field_103" at 959,515 size 33x20; Text '.2'
   TextField "Text field_104" at 959,539 size 33x20; Text '.3'
   TextField "Text field_105" at 959,563 size 33x20; Text '.4'
   TextField "Text field_106" at 959,587 size 33x20; Text '.5'
   TextField "Text field_107" at 959,611 size 33x20; Text '.6'
   TextField "Text field_108" at 959,635 size 33x20; Text '.7'
   TextField "Text field_109" at 858,467 size 33x20; Text '.0'
   TextField "Text field_110" at 858,491 size 33x20; Text '.1'
   TextField "Text field_111" at 858,515 size 33x20; Text '.2'
   TextField "Text field_112" at 858,539 size 33x20; Text '.3'
   TextField "Text field_113" at 858,563 size 33x20; Text '.4'
   TextField "Text field_114" at 858,587 size 33x20; Text '.5'
   TextField "Text field_115" at 858,611 size 33x20; Text '.6'
   TextField "Text field_116" at 858,635 size 33x20; Text '.7'
   TextField "Text field_117" at 986,467 size 33x20; Text '.0'
   TextField "Text field_118" at 986,491 size 33x20; Text '.1'
   TextField "Text field_119" at 986,515 size 33x20; Text '.2'
   TextField "Text field_120" at 986,539 size 33x20; Text '.3'
   TextField "Text field_121" at 986,563 size 33x20; Text '.4'
   TextField "Text field_122" at 986,587 size 33x20; Text '.5'
   TextField "Text field_123" at 986,611 size 33x20; Text '.6'
   TextField "Text field_124" at 986,635 size 33x20; Text '.7'
   TextField "Text field_125" at 797,447 size 43x23; Text '1'
   TextField "Text field_126" at 869,447 size 43x23; Text '3'
   TextField "Text field_127" at 925,447 size 43x23; Text '5'
   TextField "Text field_128" at 997,447 size 43x23; Text '7'
   TextField "Text field_129" at 797,225 size 43x23; Text '0'
   TextField "Text field_130" at 869,225 size 43x23; Text '2'
   TextField "Text field_131" at 925,225 size 43x23; Text '4'
   TextField "Text field_132" at 997,225 size 43x23; Text '6'
   TextField "Text field_133" at 687,447 size 43x23; Text '125'
   TextField "Text field_134" at 89,201 size 135x23; Text 'POWER SUPPLY'
   Softkey "Softkey_F1" at 0,0 size 0x0
      on KeyDown: ActivateScreen("1. MAIN", 0)
   Softkey "Softkey_F2" at 0,0 size 0x0
      on KeyDown: ActivateScreen("2. VFD 2 - 5", 0)
   Softkey "Softkey_F3" at 0,0 size 0x0
      on KeyDown: ActivateScreen("3. VFD 6 - 9", 0)
   Softkey "Softkey_F4" at 0,0 size 0x0
      on KeyDown: ActivateScreen("4. VFD 10 - 13", 0)
   Softkey "Softkey_F5" at 0,0 size 0x0
      on KeyDown: ActivateScreen("5. VFD 14 - 17", 0)
   Softkey "Softkey_F6" at 0,0 size 0x0
      on KeyDown: ActivateScreen("6. VFD 18 - 21", 0)
   Softkey "Softkey_F7" at 0,0 size 0x0
      on KeyDown: ActivateScreen("7. VFD 22 - 23", 0)
   Softkey "Softkey_F8" at 0,0 size 0x0
      on KeyDown: ActivateScreen("8. ALARM", 0)
   Softkey "Softkey_F9" at 0,0 size 0x0
      on KeyDown: ActivateScreen("9. VFD PROFIBUS", 0)
   Softkey "Softkey_F10" at 0,0 size 0x0
      on KeyDown: ActivateScreen("10. SETTINGS", 0)
*)